           // 3) SUBIDA de req_id → congelar receta. NO publicar id_ok todavía.
           IF (#SupervisorCmdReqId AND NOT #L_IdEvalDone) THEN
               #Cfg_Pns := #SupervisorCmdPns;
               #Cfg_ReferencePart := #SupervisorCmdReferencePart;
               #Cfg_EndEffector := #SupervisorCmdEndEffector;
               #Cfg_UtTeach := #SupervisorCmdUtTech;
               #Cfg_TeachReq := #SupervisorCmdTeachReq;
               #Cfg_PaCheckReq := #SupervisorCmdPaCheckReq;
               #Cfg_TcgReq := #SupervisorCmdTcgReq;

               //4) Resuelve índices de programa por pieza (tu mapeo PIEZA1/2/3)
               IF #Cfg_ReferencePart = 'RefA400M' AND #Cfg_Pns ='M551B2810006-A01' THEN
                   //PART NUMBER QUE ME ENVIARÁ DE LA PIEZA SERÁ M551B2810006-A01 
                   //  REVESTIMIENTO INF IZQ - A400M
                   #PartProgIdx := 1;
                   #RefProgIdx := 1;
               ELSIF #Cfg_ReferencePart = 'RefF10X' AND #Cfg_Pns ='F46C551713119B01'   THEN
                   //PART NUMBER QUE ME ENVIARÁ SERÁ F46C551713110B01
                   //CARENA INF. IZQ HTP/VTP - Sandwich - FALCON
                   #PartProgIdx := 2;
                   #RefProgIdx := 2;
               ELSIF #Cfg_ReferencePart = 'RefEFA' AND #Cfg_Pns ='J57462100-406' THEN
                   #PartProgIdx := 3;
                   #RefProgIdx := 3;
               ELSE
                   #PartProgIdx := 100;
                   #RefProgIdx := 100;
               END_IF;

               #L_IdEvalDone := TRUE;
           END_IF;

           // 5) BAJADA de req_id → PUBLICAR id_ok y decidir salto.
           IF ((NOT #SupervisorCmdReqId) AND #L_IdEvalDone) THEN

               //5.1) Calcula PclstatusIdOk
               #PlcStatusIdOk :=
               ("PlcStatus".plcOk AND "SupervisorCmd".supervisorOk AND "PlcStatus".robotOk AND "PlcStatus".safetyOk
               AND "PlcStatus".airOk AND "PlcStatus".inspWaterOk AND "PlcStatus".tankWaterOk)
               AND (#Cfg_EndEffector >= 1) AND (#Cfg_EndEffector <= 5);

               #PlcStatusIdRunning := FALSE;

               //5.2)Decide siguiente STEP
               IF NOT #PlcStatusIdOk THEN
                   #PlcStatusStepPlc := #cSTEP_ID;
               ELSE
                   IF #Cfg_TeachReq THEN
                       #PlcStatusStepPlc := #cSTEP_TEACH;
                   ELSE
                       #PlcStatusStepPlc := #cSTEP_STARTUS;
                   END_IF;
               END_IF;

               #L_IdEvalDone := FALSE;
           END_IF;


           // ===============================================================
           // 2) TEACHING (pág. 4) — multi-PN: rearmar teach_ready por PN
           // FÍSICO: si la herramienta necesaria para teaching no está montada,
           // el KUKA cambia en Staübli al stand indicado (usa Supervisor.end-effector).
           // Luego, el KUKA se mueve al INICIO del PN siguiente y pone un bit de “en posición”.
           // Ese bit alimenta TeachAtStart=TRUE. Entonces EL PLC arma teach_ready (p. 4).
           // Repetir por cada PN mientras teach_app_running=TRUE.
           // ===============================================================
           (*  #cSTEP_TEACH:

             IF "SupervisorCmd".teachAppRunning THEN
                   IF (NOT "SupervisorCmd".teachRunning) AND TeachAtStart THEN
                       "PlcStatus".teachReady := TRUE;
                   END_IF;

                   IF "SupervisorCmd".teachRunning THEN
                       "PlcStatus".teachReady := FALSE;
                       teachWasRunning := TRUE;
                   END_IF;

                   // Fin de una trayectoria de teaching (sin abandonar la app)
                   IF (NOT "SupervisorCmd".teachRunning) AND teachWasRunning THEN
                       teachWasRunning := FALSE;
                   END_IF;

               ELSE
                   // Cierre de la app: salto según teach_state
                   IF "SupervisorCmd".teachState THEN
                       "PlcStatus".stepPlc := cSTEP_STARTUS;
                   ELSE
                       "PlcStatus".stepPlc := cSTEP_ID;
                   END_IF;
               END_IF;
           END_IF;*)




           // ===============================================================
           // 3) START US (pág. 5) — armar cuando “previous task done”
           // FÍSICO: KUKA AUT EXT cambia (si hace falta) al efector de INSPECCIÓN
           // requerido (Supervisor.end-effector, p. 1). Cuando:
           //   - Herramienta correcta acoplada (Staübli OK),
           //   - servicios/enclavamientos OK (safety/air/water/tank),
           //   - robot en posición segura para inicializar el UT,
           // el secuenciador pone StartUSReady=TRUE. El PLC arma start_us_ready.
           // Supervisor hace init UT (start_us_running/state_us). (p. 5)
           // ===============================================================
       #cSTEP_STARTUS:

           // Al entrar, ordena al robot cargar la herramienta decidida en ID
           IF #firstScan THEN
               #SupervisorCmdSeq := #SupervisorCmdSeq + 1;
               #WantCode_uint := #cKUKA_REQ_TOOL;
               #WantToolRequestId := (#Cfg_EndEffector);       // 1..5
           END_IF;

           // El PLC arma startUsReady SI el entorno/robot están listos y todavía no corre
           IF #StartUSReady AND (#WantCode_uint = 0) AND ("ToolInRobot_DB".toolInRobot_Num = #Cfg_EndEffector) AND NOT #SupervisorCmdStartUsRunning THEN
               #PlcStatusStartUsReady := TRUE;
           END_IF;

           // Cuando arranca, baja el "ready" y registra que realmente empezó
           IF #SupervisorCmdStartUsRunning THEN
               #PlcStatusStartUsReady := FALSE;
               #startUSWasRunning := TRUE;
           END_IF;

           // Al terminar: salto a PA o a Gain según lo congelado en ID
           IF (NOT #SupervisorCmdStartUsRunning)  AND #startUSWasRunning THEN
               #startUSWasRunning := FALSE;
               IF NOT #SupervisorCmdStateUs THEN
                   #PlcStatusStepPlc := #cSTEP_ID;
               ELSE
                   IF #Cfg_PaCheckReq THEN
                       #PlcStatusStepPlc := #cSTEP_PA_BAL;
                   ELSE
                       #PlcStatusStepPlc := #cSTEP_GAIN;
                   END_IF;
               END_IF;
           END_IF;


           // ===============================================================
           // 4) DEAD ELEMENT CHECK & BALANCING (pág. 6)
           //FÍSICO: KUKA va a la pieza Perspex de calibración y, cuando está en
           // [CORREGIDO] Lógica secuencial robusta, GOTO determinista y Retracción.
           // ===============================================================
       #cSTEP_PA_BAL:
           CASE #paBalSubStep OF
               0: // Inicialización y GOTO_PERSPEX
                   // [MEJORA] Siempre enviar comando GOTO en firstScan.
                   IF #firstScan THEN
                       #SupervisorCmdSeq := #SupervisorCmdSeq + 1;
                       #WantCode_uint := #cKUKA_GOTO_PERSPEX;
                   END_IF;
                   #paBalSubStep := 10;
               10: // Esperar Posición en Perspex     
                   // [MEJORA] Esperar posición Y canal libre (Race condition fix)
                   IF #kukaAtPerspexPos AND (#WantCode_uint = 0) THEN
                       #paBalSubStep := 20;
                   END_IF;
               20: // Ready for Dead Element Check     
                   IF NOT "SupervisorCmd".elemRunning THEN
                       "PlcStatus".paCheckReady := TRUE;
                   END_IF;
                   IF "SupervisorCmd".elemRunning THEN
                       "PlcStatus".paCheckReady := FALSE;
                       #paBalSubStep := 30;
                   END_IF;
               30: // Dead Element Check Running       
                   IF NOT "SupervisorCmd".elemRunning THEN
                       IF "SupervisorCmd".elemState THEN
                           #paBalSubStep := 40; // OK -> Balancing
                       ELSE
                           // KO -> Almacenar resultado y retraer
                           #tempNextStep := #cSTEP_ID;
                           #paBalSubStep := 60; // Ir a retracción
                       END_IF;
                   END_IF;
               40: // Ready for Balancing (Supervisor inicia automáticamente)        
                   IF "SupervisorCmd".balRunning THEN
                       #paBalSubStep := 50;
                   END_IF;
               50: // Balancing Running        
                   IF NOT "SupervisorCmd".balRunning THEN
                       // Determinar el siguiente paso
                       IF "SupervisorCmd".balState THEN
                           #tempNextStep := #cSTEP_GAIN; // OK
                       ELSE
                           #tempNextStep := #cSTEP_ID; // KO
                       END_IF;
                       #paBalSubStep := 60; // Proceder a retracción
                   END_IF;

                   // --- [MEJORA] LÓGICA DE RETRACCIÓN ESPECÍFICA ---
               60: // Ordenar RETRACT_PERSPEX
                   // [MEJORA] Esperar disponibilidad del despachador (Race condition fix)
                   IF (#WantCode_uint = 0) THEN
                       #SupervisorCmdSeq := #SupervisorCmdSeq + 1;
                       #WantCode_uint := #cKUKA_RETRACT_PERSPEX; // 101
                       #paBalSubStep := 70;
                   END_IF;

               70: // Esperar Fin de Retracción
                   // Robot terminó (WantCode_uint reseteado por el despachador)
                   IF (#WantCode_uint = 0) THEN
                       // Transición al paso almacenado
                       "PlcStatus".stepPlc := #tempNextStep;
                   END_IF;
           END_CASE;

           // ===============================================================
           // 5) GAIN ADJUSTMENT (pág. 7)
           // FÍSICO: KUKA se posiciona en la referencia para ganancia estática;
           // [CORREGIDO] Lógica secuencial robusta, GOTO determinista y Retracción.
           // ===============================================================
       #cSTEP_GAIN:

           CASE #gainSubStep OF
               0: // Inicialización y GOTO_GAIN
                   // [MEJORA] Siempre enviar comando GOTO en firstScan.
                   IF #firstScan THEN
                       #SupervisorCmdSeq := #SupervisorCmdSeq + 1;
                       #WantCode_uint := #cKUKA_GOTO_GAIN;
                   END_IF;
                   #gainSubStep := 10;

               10: // Esperar Posición en Gain    
                   // [MEJORA] Esperar posición Y canal libre (Race condition fix)
                   IF #kukaAtGainPos AND (#WantCode_uint = 0) THEN
                       #gainSubStep := 20;
                   END_IF;

               20: // Ready for Gain (Supervisor)    
                   IF NOT "SupervisorCmd".gainRunning THEN
                       "PlcStatus".gainReady := TRUE;
                   END_IF;

                   IF "SupervisorCmd".gainRunning THEN
                       "PlcStatus".gainReady := FALSE;
                       #gainSubStep := 30;
                   END_IF;

               30: // Gain Running
                   IF NOT "SupervisorCmd".gainRunning THEN
                       // Determinar siguiente paso
                       IF "SupervisorCmd".gainState THEN
                           IF #Cfg_TcgReq THEN
                               #tempNextStep := #cSTEP_TCG;
                           ELSE
                               #tempNextStep := #cSTEP_SCAN_REF;
                           END_IF;
                       ELSE
                           #tempNextStep := #cSTEP_ID; // KO        
                       END_IF;
                       #gainSubStep := 40; // Proceder a retracción
                   END_IF;

                   // --- [MEJORA] LÓGICA DE RETRACCIÓN ESPECÍFICA ---
               40: // Ordenar RETRACT_GAIN
                   // [MEJORA] Esperar disponibilidad del despachador (Race condition fix) 
                   IF (#WantCode_uint = 0) THEN
                       #SupervisorCmdSeq := #SupervisorCmdSeq + 1;
                       #WantCode_uint := #cKUKA_RETRACT_GAIN; // 102
                       #gainSubStep := 50;
                   END_IF;
               50: // Esperar Fin de Retracción         
                   IF (#WantCode_uint = 0) THEN
                       "PlcStatus".stepPlc := #tempNextStep;
                   END_IF;

           END_CASE;




           // ===============================================================
           // (6) TCG CHECK / ADJUSTMENT — pág. 8 (multiposición)
           // FÍSICO: KUKA recorre varias posiciones TCG. Para cada posición:
           // [CORREGIDO] Handshake Manager, GOTO determinista, Race Condition Fix y Retracción.
           // ===============================================================
       #cSTEP_TCG:

           // [MEJORA] Siempre ordenar el primer movimiento al entrar.    
           IF #firstScan THEN
               #SupervisorCmdSeq := #SupervisorCmdSeq + 1;
               #WantCode_uint := #cKUKA_GOTO_TCG;
               #WantIndex := (#tcgIndex); // Debería ser 1
               #waitingNextTCGPos := TRUE;
           END_IF;

           // Rearme de espera.
           // [MEJORA] Esperar a KUKA en posición Y que el canal esté libre (Race condition fix).
           IF #waitingNextTCGPos AND #kukaAtTCGPos AND (#WantCode_uint = 0) THEN
               #waitingNextTCGPos := FALSE;
           END_IF;

           // tcg_ready sólo si no mide, no esperamos pos, y el Handshake Manager está libre.
           IF (NOT "SupervisorCmd".tcgInProgress) AND (NOT #waitingNextTCGPos) AND (#handshakeStep = 0) THEN
               "PlcStatus".tcgReady := TRUE;
           ELSE
               // Asegurar que tcgReady baja si alguna condición falla (ej. Supervisor inicia medición)     
               "PlcStatus".tcgReady := FALSE;
           END_IF;

           // --- [MEJORA] Handshake Manager (4-way Acknowledge) - PDF Pág. 8 ---
           CASE #handshakeStep OF
               0: // IDLE: Esperar solicitud (Priorizadas)
                   // Solo aceptar si no estamos esperando movimiento ni midiendo
                   IF (NOT #waitingNextTCGPos) AND (NOT "SupervisorCmd".tcgInProgress) THEN
                       IF "SupervisorCmd".tcgNextStep THEN
                           #handshakeStep := 1; // NEXT
                       ELSIF "SupervisorCmd".reqRefPart THEN
                           #handshakeStep := 2; // ReqRefPart (Salida)
                       ELSIF "SupervisorCmd".reqStopCycle THEN
                           #handshakeStep := 3; // StopCycle (Salida)
                       ELSIF "SupervisorCmd".reqTcgAdj THEN
                           #handshakeStep := 4; // TcgAdj (Permanece en TCG) 
                       END_IF;
                   END_IF;

                   //1, 2, 3, 4: // SOLICITUD RECIBIDA: Enviar Acknowledge     
                   "PlcStatus".acknowledge := TRUE;
                   #handshakeStep := #handshakeStep + 10; // Pasar a esperar bajada
                   // --- Esperar Bajada de Solicitud ---    
               11: // NEXT    
                   IF NOT "SupervisorCmd".tcgNextStep THEN
                       "PlcStatus".acknowledge := FALSE;
                       // Acción NEXT: Pasar a esperar disponibilidad del canal antes de enviar.
                       #handshakeStep := 21;
                   END_IF;
               12: // ReqRefPart (Salida)
                   IF NOT "SupervisorCmd".reqRefPart THEN
                       "PlcStatus".acknowledge := FALSE;
                       // Acción: Preparar retracción antes de saltar.
                       #tempNextStep := #cSTEP_SCAN_REF;
                       #handshakeStep := 50; // Ir a retracción
                   END_IF;

               13: // StopCycle (Salida)     
                   IF NOT "SupervisorCmd".reqStopCycle THEN
                       "PlcStatus".acknowledge := FALSE;
                       // Acción: Preparar retracción antes de saltar. 
                       #tempNextStep := #cSTEP_ID;
                       #handshakeStep := 50; // Ir a retracción
                   END_IF;

               14: // TcgAdj (Permanece)     
                   IF NOT "SupervisorCmd".reqTcgAdj THEN
                       "PlcStatus".acknowledge := FALSE;
                       // Acción: Permanecer en TCG (Modo Ajuste).   
                       #handshakeStep := 0;
                   END_IF;

                   // --- Ejecución de NEXT (Sincronización con Despachador) ---
               21: // EJECUTAR NEXT (Wait for Dispatcher)
                   // [MEJORA] Evitar condición de carrera del despachador.
                   IF (#WantCode_uint = 0) THEN
                       // Canal libre -> Enviar comando GOTO_TCG
                       #tcgIndex := #tcgIndex + 1;
                       #SupervisorCmdSeq := #SupervisorCmdSeq + 1;
                       #WantCode_uint := #cKUKA_GOTO_TCG;
                       #WantIndex := (#tcgIndex);
                       #waitingNextTCGPos := TRUE;
                       #handshakeStep := 0;
                   END_IF;

                   // --- LÓGICA DE RETRACCIÓN ESPECÍFICA (Para salidas del paso TCG) ---        
               50: // Ordenar RETRACT_TCG
                   IF (#WantCode_uint = 0) THEN
                       #SupervisorCmdSeq := #SupervisorCmdSeq + 1;
                       #WantCode_uint := #cKUKA_RETRACT_TCG; // 103
                       #handshakeStep := 60;
                   END_IF;

               60: // Esperar Fin de Retracción      
                   IF (#WantCode_uint = 0) THEN
                       "PlcStatus".stepPlc := #tempNextStep; // Ir al paso almacenado
                       #handshakeStep := 0;
                   END_IF;
           END_CASE;



           // ===============================================================
           // (7) SCAN REFERENCE ACQUISITION — pág. 10
           // FÍSICO: KUKA carga PN/frame y se coloca en el punto de INICIO de
           // la trayectoria de referencia. Tu lógica pone AtRefScanStart=TRUE cuando
           // está en posición. 
           // // [MEJORA] GOTO determinista y Sincronización robusta.
           // ===============================================================
       #cSTEP_SCAN_REF:

           // Validación mínima de parámetros de scan que el PLC publica al Supervisor
           #validScanParams := (LEN("PlcStatus".idScan) > 0) AND ("PlcStatus".xSize > 0.0) AND ("PlcStatus".ySize > 0.0);

           // [MEJORA] Siempre enviar comando GOTO en firstScan.
           IF #firstScan THEN
               #SupervisorCmdSeq := #SupervisorCmdSeq + 1;
               #WantCode_uint := #cKUKA_GOTO_REF_START; // CASE 420
               #WantProgRequestId := (#RefProgIdx); // índice de programa REF por pieza
           END_IF;

           // Permiso de arranque
           // [MEJORA] Esperar posición Y canal libre antes de dar Ready.
           IF #kukaAtRefScanStartPos AND (#WantCode_uint = 0) AND #validScanParams AND NOT "SupervisorCmd".scanRefRunning THEN
               "PlcStatus".scanRefStart := TRUE;
           END_IF;

           // Cuando el Supervisor arranca → ejecutar trayectoria (CASE 432)
           IF (NOT #scanRefWasRunning) AND "SupervisorCmd".scanRefRunning THEN
               // [MEJORA] Esperar a que el despachador esté libre antes de enviar RUN.
               IF (#WantCode_uint = 0) THEN
                   #SupervisorCmdSeq := #SupervisorCmdSeq + 1;
                   #WantCode_uint := #cKUKA_RUN_REF_PATH;
                   #WantProgRequestId := (#RefProgIdx);
                   #scanRefWasRunning := TRUE; // Marcar como iniciado solo tras enviar comando
               END_IF;
           END_IF;

           IF "SupervisorCmd".scanRefRunning THEN
               // Bajar Ready cuando el robot termina físicamente  
               IF #kukaRefScanFinished THEN
                   "PlcStatus".scanRefStart := FALSE;
               END_IF;
           END_IF;

           // Fin del escaneo    
           IF (NOT "SupervisorCmd".scanRefRunning) AND #scanRefWasRunning THEN
               #scanRefWasRunning := FALSE;
               "PlcStatus".scanRefStart := FALSE;
               IF NOT "SupervisorCmd".scanRefState THEN
                   "PlcStatus".stepPlc := #cSTEP_ID;
               ELSE
                   "PlcStatus".stepPlc := #cSTEP_SCAN_INSP;
               END_IF;
           END_IF;


           // ===============================================================
           // (8) SCAN INSPECTION — pág. 11
           // FÍSICO: KUKA se coloca en INICIO de la(s) trayectoria(s) de inspección
           // [CORREGIDO] Handshake Manager, GOTO determinista y Sincronización robusta.
           // ===============================================================
       #cSTEP_SCAN_INSP:

           #validScanParams := (LEN("PlcStatus".idScan) > 0) AND ("PlcStatus".xSize > 0.0) AND ("PlcStatus".ySize > 0.0);

           // [MEJORA] Siempre enviar comando GOTO en firstScan.
           IF #firstScan THEN
               #SupervisorCmdSeq := #SupervisorCmdSeq + 1;
               #WantCode_uint := #cKUKA_GOTO_INSP_START;
               #WantProgRequestId := (#PartProgIdx);
           END_IF;

           // Permiso de arranque
           // [MEJORA] Esperar posición, canal libre y handshake libre antes de dar Ready.
           IF #kukaAtInspScanStartPos AND (#WantCode_uint = 0) AND #validScanParams AND NOT "SupervisorCmd".scanInsprunning AND (#handshakeStep = 0) THEN
               "PlcStatus".scanInspStart := TRUE;
           END_IF;

           // Al arrancar → ejecutar trayectoria (CASE 433)
           IF (NOT #scanInspWasRunning) AND "SupervisorCmd".scanInsprunning THEN
               // [MEJORA] Esperar a que el despachador esté libre antes de enviar RUN.
               IF (#WantCode_uint = 0) THEN
                   #SupervisorCmdSeq := #SupervisorCmdSeq + 1;
                   #WantCode_uint := #cKUKA_RUN_INSP_PATH;
                   #WantProgRequestId := (#PartProgIdx);
                   #scanInspWasRunning := TRUE; // Marcar como iniciado solo tras enviar comando
               END_IF;
           END_IF;


           IF "SupervisorCmd".scanInsprunning THEN
               // Bajar Ready cuando el robot termina físicamente
               IF #kukaInspScanFinished THEN
                   "PlcStatus".scanInspStart := FALSE;
               END_IF;
           END_IF;

           // Fin del escaneo 
           IF (NOT "SupervisorCmd".scanInsprunning) AND #scanInspWasRunning THEN
               #scanInspWasRunning := FALSE;
               "PlcStatus".scanInspStart := FALSE;

               IF NOT "SupervisorCmd".scanInspState THEN
                   "PlcStatus".stepPlc := #cSTEP_ID;
               ELSE
                   // Escaneo OK -> Activar Handshake Manager para esperar req_verif
                   #handshakeStep := 1;
               END_IF;
           END_IF;
           // [MEJORA] Handshake Manager (4-way) para req_verif (PDF Pág. 11)     
               CASE #handshakeStep OF
                   1: // Esperando req_verif
                       IF "SupervisorCmd".reqVerif THEN
                           #handshakeStep := 2;
                       END_IF;

                   2: // Enviar Acknowledge       
                       "PlcStatus".acknowledge := TRUE;
                       #handshakeStep := 3;

                   3: // Esperar bajada de req_verif    
                       IF NOT "SupervisorCmd".reqVerif THEN
                           "PlcStatus".acknowledge := FALSE;
                           // Acción: Saltar a Verificación 
                           "PlcStatus".stepPlc := #cSTEP_SCAN_REF_VERIF;
                           #handshakeStep := 0;
                       END_IF;
               END_CASE;





           // ===============================================================
           // (9) SCAN REFERENCE VERIFICATION — pág. 12
           // FÍSICO: KUKA vuelve al INICIO de la trayectoria de verificación de ref.
           // [CORREGIDO] Handshake Manager, Orden Faltante, GOTO y Sincronización.
           // ===============================================================
       #cSTEP_SCAN_REF_VERIF:

           #validScanParams := (LEN("PlcStatus".idScan) > 0) AND ("PlcStatus".xSize > 0.0) AND ("PlcStatus".ySize > 0.0);

           // [MEJORA] Siempre enviar comando GOTO en firstScan.
           IF #firstScan THEN
               #SupervisorCmdSeq := #SupervisorCmdSeq + 1;
               #WantCode_uint := #cKUKA_GOTO_REF_START;
               #WantProgRequestId := (#RefProgIdx);
           END_IF;
           // Permiso de arranque    
           // [MEJORA] Esperar posición, canal libre y handshake libre antes de dar Ready.
           IF #kukaAtRefScanStartPos AND (#WantCode_uint = 0) AND #validScanParams AND NOT "SupervisorCmd".scanRefRunning AND (#handshakeStep = 0) THEN
               "PlcStatus".scanRefStart := TRUE;
           END_IF;

           // [CORRECCIÓN] Al arrancar -> ejecutar trayectoria (Faltaba esta orden)
           IF (NOT #scanRefWasRunning) AND "SupervisorCmd".scanRefRunning THEN
               // [MEJORA] Esperar a que el despachador esté libre antes de enviar RUN.
               IF (#WantCode_uint = 0) THEN
                   #SupervisorCmdSeq := #SupervisorCmdSeq + 1;
                   #WantCode_uint := #cKUKA_RUN_REF_PATH; // 432
                   #WantProgRequestId := (#RefProgIdx);
                   #scanRefWasRunning := TRUE; // Marcar como iniciado solo tras enviar comando
               END_IF;
           END_IF;

           IF "SupervisorCmd".scanRefRunning THEN
               // [CORRECCIÓN] Bajar scanRefStart cuando el robot termina (PDF p.12).
               IF #kukaRefScanFinished THEN
                   "PlcStatus".scanRefStart := FALSE;
               END_IF;
           END_IF;

           // Fin del escaneo de verificación
           IF (NOT "SupervisorCmd".scanRefRunning) AND #scanRefWasRunning THEN
               #scanRefWasRunning := FALSE;
               "PlcStatus".scanRefStart := FALSE;
               IF NOT "SupervisorCmd".scanRefState THEN
                   "PlcStatus".stepPlc := #cSTEP_ID;
               ELSE
                   // OK -> Activar Handshake Manager para esperar decisiones    
                   #handshakeStep := 1;
               END_IF;
           END_IF;

           // [MEJORA] Handshake Manager (4-way) (PDF Pág. 12)
           CASE #handshakeStep OF
               1: // Esperando decisiones (Priorizadas)
                   IF "SupervisorCmd".reqPreEval THEN
                       #handshakeStep := 2; // Pre-eval
                   ELSIF "SupervisorCmd".reqIdentificationState THEN
                       #handshakeStep := 3; // Nuevo ciclo
                   END_IF;
                   // 2, 3: // Enviar Acknowledge
                   "PlcStatus".acknowledge := TRUE;
                   #handshakeStep := #handshakeStep + 10;
               12: // Esperar bajada (Pre-eval)     
                   IF NOT "SupervisorCmd".reqPreEval THEN
                       "PlcStatus".acknowledge := FALSE;
                       "PlcStatus".stepPlc := #cSTEP_PRE_EVAL;
                       #handshakeStep := 0;
                   END_IF;

               13: // Esperar bajada (Nuevo Ciclo)      
                   IF NOT "SupervisorCmd".reqIdentificationState THEN
                       "PlcStatus".acknowledge := FALSE;
                       // Nota: No se requiere GOTO_SAFE aquí, ya que el escaneo no es peligroso.
                       "PlcStatus".stepPlc := #cSTEP_ID;
                       #handshakeStep := 0;
                   END_IF;
           END_CASE;

           // ===============================================================
           // (10) PRE‑EVALUATION / MARKING — pág. 13
           // FÍSICO: si la herramienta de marcado no está montada, el KUKA cambia
           // en Staübli al stand de “marking” según requiera el proceso; tras estar
           // [CORREGIDO] Gestión de herramienta, ejecución física, Handshake y movimiento seguro.
           // ===============================================================
       #cSTEP_PRE_EVAL:

           // --- [MEJORA] Handshake Manager (4-way) para Nuevo ciclo + GOTO_SAFE ---  
           CASE #handshakeStep OF
               0: // Idle: Esperar solicitud de nuevo ciclo       
                   // Solo permitir si el marcado no está en curso   
                   IF "SupervisorCmd".reqIdentificationState AND (NOT "PlcStatus".markRunning) THEN
                       #handshakeStep := 1;
                   END_IF;
               1: // Enviar Ack    
                   "PlcStatus".acknowledge := TRUE;
                   #handshakeStep := 2;
               2: // Esperar bajada de la solicitud
                   IF NOT "SupervisorCmd".reqIdentificationState THEN
                       "PlcStatus".acknowledge := FALSE;
                       // Acción: Preparar para ir a Safe antes de ID    
                       #handshakeStep := 3;
                   END_IF;

                   // [MEJORA] Mover a Safe antes de saltar a ID      
               3: // Enviar GOTO_SAFE (Esperar disponibilidad del despachador)   
                   IF (#WantCode_uint = 0) THEN
                       #SupervisorCmdSeq := #SupervisorCmdSeq + 1;
                       //#WantCode_uint := #cKUKA_GOTO_SAFE; // 100
                       #handshakeStep := 4;
                   END_IF;

               4: // Esperar fin de GOTO_SAFE
                   IF (#WantCode_uint = 0) THEN
                       // Llegó a Safe -> Saltar a ID
                       "PlcStatus".stepPlc := #cSTEP_ID;
                       #handshakeStep := 0;
                   END_IF;
           END_CASE;

           // --- [MEJORA] Máquina de estados de Marcado ---
           CASE #markingSubStep OF
               0: // Inicialización (Al entrar al paso)
                   #markingSubStep := 10;
               10: // Cambio de Herramienta (a Marcador)     
                   // Solo si no la tiene ya y los canales están libres
                   IF ("ToolInRobot_DB".toolInRobot_Num <> 3) AND (#WantCode_uint = 0) AND (#handshakeStep = 0) THEN
                       #SupervisorCmdSeq := #SupervisorCmdSeq + 1;
                       #WantCode_uint := #cKUKA_REQ_TOOL;
                       #WantToolRequestId := #cTOOL_MARKER;
                   END_IF;

                   // Transición cuando tenga la herramienta y el canal esté libre    
                   IF ("ToolInRobot_DB".toolInRobot_Num = #cTOOL_MARKER) AND (#WantCode_uint = 0) THEN
                       #markingSubStep := 20;
                   END_IF;

               20: // Esperar Petición de Marcado (reqMark)
                   // Solo si el handshake general está libre
                   IF "SupervisorCmd".reqMark AND (#handshakeStep = 0) THEN
                       // 1. Transferir coordenadas al buffer (Asume Supervisor.pointCoordinates es ARRAY[0..5] OF REAL)
                       // #WantMarkCoords[0] := "SupervisorCmd".pointCoordinates[0]; // X
                       // ... (Copiar Y, Z, A, B, C) ...
                       // 2. Preparar estado y pasar a envío de comando
                       "PlcStatus".markState := FALSE;
                       "PlcStatus".markRunning := TRUE;
                       #markingSubStep := 30;
                   END_IF;

               30: // Enviar Comando al Robot (Esperar disponibilidad)    
                   // [MEJORA] Esperar a que el despachador esté libre.
                   IF (#WantCode_uint = 0) THEN
                       #SupervisorCmdSeq := #SupervisorCmdSeq + 1;
                       #WantCode_uint := #cKUKA_MARK_POINT; // Código 501
                       #markingSubStep := 40;
                   END_IF;

               40: // Ejecución en Progreso (Esperar fin en KUKA)  
                   // Esperar a que el robot termine el comando (WantCode_uint vuelve a 0)
                   IF (#WantCode_uint = 0) THEN
                       // El marcado ha terminado físicamente.
                       "PlcStatus".markState := #MarkingDone; // Leer resultado físico
                       #markingSubStep := 50;
                   END_IF;

               50: // Finalizado (Esperar que Supervisor baje reqMark - PDF p.13)
                   IF NOT "SupervisorCmd".reqMark THEN
                       "PlcStatus".markRunning := FALSE;
                       "PlcStatus".markRunning := FALSE;
                   END_IF;

           END_CASE;
       ELSE
           "PlcStatus".stepPlc := #cSTEP_ID;

   END_CASE;


   // ---------------------------------------------------------------
   // [2] DESPACHO AL KUKA (toggle goTrigger cuando el canal esté libre)
   //     • Este bloque “consume” el slot WantCmd → publica parámetros
   //       en los registros PNIO (con SWAP) → toggle de goTrigger.
   //     • El robot deberá igualar rbDone := goTrigger al terminar.
   // ---------------------------------------------------------------

   CASE #state OF
       0: // IDLE -> GO == ACK

           // "cancelGo" := FALSE;

           IF (#SupervisorCmdSeq <> #lastSeq) THEN

               IF  "goTrigger" = "rbDone" THEN

                   #code_int := #WantCode_uint;  // “code_int” que viajará al KRC

                   // (Códigos existentes 201, 414, 420, 432, 421, 433 se mantienen igual)

                   IF #code_int = 201 THEN
                       // id de herramienta → WORD+SWAP
                       // #Cfg_EndEffector
                       #toolReqId := SWAP(INT_TO_WORD(#WantToolRequestId));

                   END_IF;

                   IF #code_int = 414 THEN  //GOTO_TCG
                       // id de herramienta → WORD+SWAP
                       "requestIndexKuka" := SWAP(UINT_TO_WORD(#WantIndex));

                   END_IF;

                   IF #code_int = 420 THEN // GOTO_REF_START
                       // id de herramienta → WORD+SWAP
                       "programReqId" := SWAP(UINT_TO_WORD(#WantProgRequestId));

                   END_IF;

                   IF #code_int = 432 THEN // RUN_REF_PATH
                       // id de herramienta → WORD+SWAP
                       "programReqId" := SWAP(UINT_TO_WORD(#WantProgRequestId));

                   END_IF;

                   IF #code_int = 421 THEN // GOTO_REF_START
                       // id de herramienta → WORD+SWAP
                       "programReqId" := SWAP(UINT_TO_WORD(#WantProgRequestId));

                   END_IF;

                   IF #code_int = 433 THEN // RUN_INSP_PATH

                       "programReqId" := SWAP(UINT_TO_WORD(#WantProgRequestId));

                   END_IF;

                   // [MEJORA] Transferencia de Coordenadas para Marcado (501)
                  // IF #code_int = #cKUKA_MARK_POINT THEN
                        // Convertir REAL a DWORD/DINT y hacer SWAP para enviar por Profinet
                        //  // Ejemplo: "ProfinetOutputs".MarkX := SWAP(REAL_TO_DWORD(#WantMarkCoords[0]));
                   //END_IF;

                   // 2) Publicar código de movimiento
                   #moveCodeKuka := SWAP(UINT_TO_WORD(#code_int));   // KRC leerá "MoveCode" = INT

                   // 3) Disparo del GO: toggle de goTrigger (rbDone ≠ goTrigger → pedido activo)
                   "goTrigger" := NOT "goTrigger";

                   #lastSeq := #SupervisorCmdSeq;          // <-- memoriza!
                   #state := 20;

               END_IF;
           END_IF;

       20: // BUSY

           //#code_int := #KukaControlCmdCode;

           // CANCEL pedido en BUSY → avisar al KRC y ACK de la ORDEN ACTIVA
           IF #code_int = 903 THEN
               "cancelGo" := TRUE;
           END_IF;

           // Fin normal (o tras el cancel, cuando KRC cierra el canal por nivel)

           IF ("rbDone" = "goTrigger") THEN
               // 4) Vaciar slot de pendiente
               #WantCode_uint := 0;
               #WantProgRequestId := 0;
               #WantToolRequestId := 0;
               #WantIndex := 0;
               #state := 0;                            // vuelve a IDLE
           END_IF;

   END_CASE;
END_REGION
END_FUNCTION_BLOCK

ORGANIZATION_BLOCK "Main"   // OB1, LAD, ProgramCycle
TITLE = "Main Program Sweep (Cycle)"
{ S7_Optimized_Access := 'TRUE' }
VERSION : 0.1
   VAR_INPUT
      Initial_Call : Bool;   // Initial call of this OB
      Remanence : Bool;   // =True, if remanent data are available
   END_VAR
   VAR_TEMP
      evtEnterSrv : Bool;   // // Eventos de modo service jog
      evtEnterAuto : Bool;   // // Eventos de modo auto
      muxSelStb : Bool;
      muxStartStb : Bool;
      muxPgno : Byte;
      u : UDInt;
   END_VAR
BEGIN

REGION Network 1 (SCL): // ====================== REANUDAR MOVIMIENTO AUTOMATICO EXTERNO ======================
   // // —— Enlaza estos símbolos a tus %I en el árbol de dispositivos ——
   //   // EStop_DI, SafeDoor_DI, AirPressure_DI, WaterInsp_DI, WaterTank_DI, RobotReady_DI, ...
   "$MOVE_ENABLE" := TRUE;
   "$I_O_ACT" := TRUE;
   //"$DRIVES_OFF" := FALSE;

   "PlcStatus".systemArmed := FALSE;
   "PlcStatus".robotInAutExt := "$EXT";
   "PlcStatus".robotInHome := "$IN_HOME";
END_REGION

REGION Network 2: REANUDAR MOVIMIENTO EN KUKA
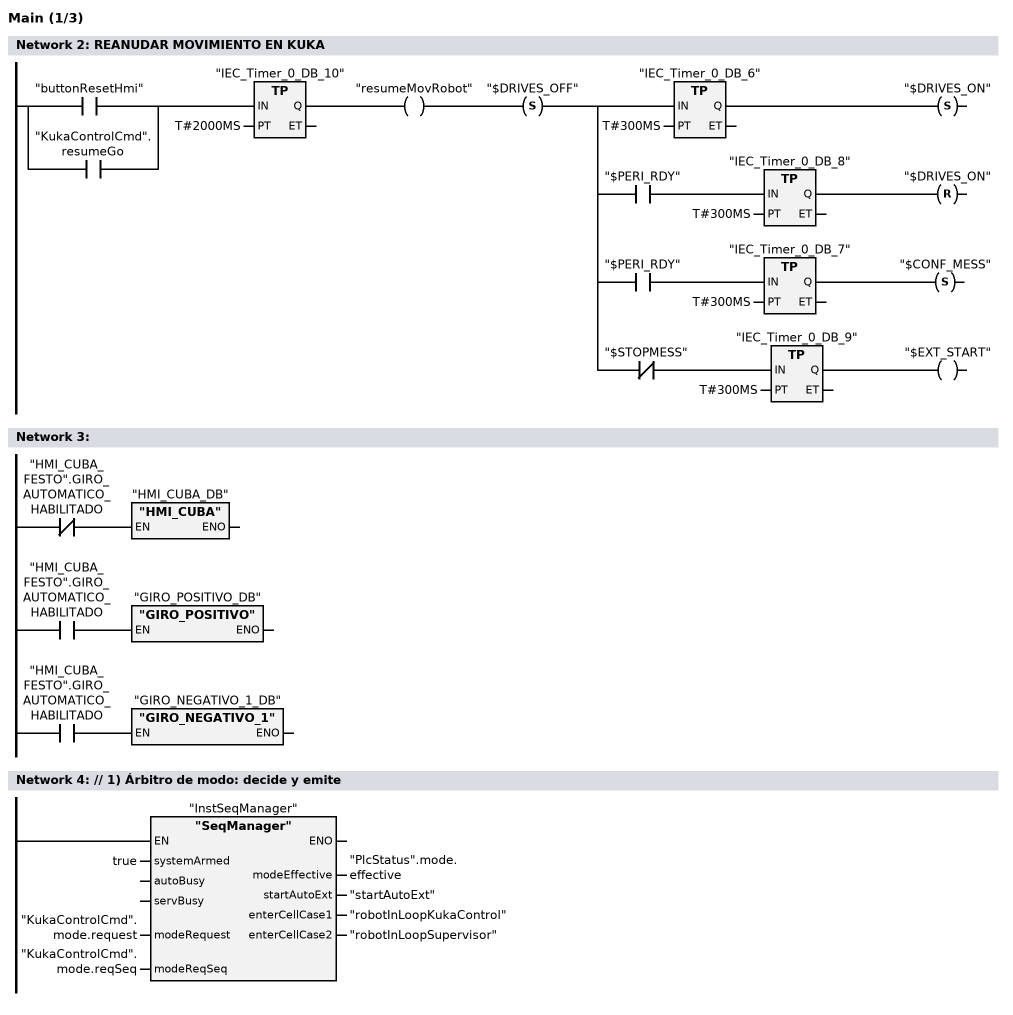
   "IEC_Timer_0_DB_10".TP(IN := "buttonResetHmi" OR "KukaControlCmd".resumeGo, PT := T#2000MS);
   "resumeMovRobot" := "IEC_Timer_0_DB_10".Q;
   IF "IEC_Timer_0_DB_10".Q THEN "$DRIVES_OFF" := TRUE; END_IF;
   "IEC_Timer_0_DB_6".TP(IN := "IEC_Timer_0_DB_10".Q, PT := T#300MS);
   IF "IEC_Timer_0_DB_6".Q THEN "$DRIVES_ON" := TRUE; END_IF;
   "IEC_Timer_0_DB_8".TP(IN := "IEC_Timer_0_DB_10".Q AND "$PERI_RDY", PT := T#300MS);
   IF "IEC_Timer_0_DB_8".Q THEN "$DRIVES_ON" := FALSE; END_IF;
   "IEC_Timer_0_DB_7".TP(IN := "IEC_Timer_0_DB_10".Q AND "$PERI_RDY", PT := T#300MS);
   IF "IEC_Timer_0_DB_7".Q THEN "$CONF_MESS" := TRUE; END_IF;
   "IEC_Timer_0_DB_9".TP(IN := "IEC_Timer_0_DB_10".Q AND NOT "$STOPMESS", PT := T#300MS);
   "$EXT_START" := "IEC_Timer_0_DB_9".Q;
END_REGION

REGION Network 3
   RUNG wire#powerrail
      I_Contact( "HMI_CUBA_FESTO".GIRO_AUTOMATICO_HABILITADO )
      "HMI_CUBA_DB"()
   END_RUNG
   RUNG wire#powerrail
      Contact( "HMI_CUBA_FESTO".GIRO_AUTOMATICO_HABILITADO )
      "GIRO_POSITIVO_DB"()
   END_RUNG
   RUNG wire#powerrail
      Contact( "HMI_CUBA_FESTO".GIRO_AUTOMATICO_HABILITADO )
      "GIRO_NEGATIVO_1_DB"()
   END_RUNG
   // the same network as SCL:
   IF NOT "HMI_CUBA_FESTO".GIRO_AUTOMATICO_HABILITADO THEN
       "HMI_CUBA_DB"();   // "HMI_CUBA"
   END_IF;
   IF "HMI_CUBA_FESTO".GIRO_AUTOMATICO_HABILITADO THEN
       "GIRO_POSITIVO_DB"();   // "GIRO_POSITIVO"
   END_IF;
   IF "HMI_CUBA_FESTO".GIRO_AUTOMATICO_HABILITADO THEN
       "GIRO_NEGATIVO_1_DB"();   // "GIRO_NEGATIVO_1"
   END_IF;
END_REGION

REGION Network 4: // 1) Árbitro de modo: decide y emite
   RUNG wire#powerrail
      "InstSeqManager"(systemArmed := true, autoBusy :=, servBusy :=, modeRequest := "KukaControlCmd".mode.request, modeReqSeq := "KukaControlCmd".mode.reqSeq, modeEffective => "PlcStatus".mode.effective, startAutoExt => "startAutoExt", enterCellCase1 => "robotInLoopKukaControl", enterCellCase2 => "robotInLoopSupervisor")
   END_RUNG
   // the same network as SCL:
   "InstSeqManager"(systemArmed := true,   // "SeqManager"
                    modeRequest := "KukaControlCmd".mode.request,
                    modeReqSeq := "KukaControlCmd".mode.reqSeq,
                    modeEffective => "PlcStatus".mode.effective,
                    startAutoExt => "startAutoExt",
                    enterCellCase1 => "robotInLoopKukaControl",
                    enterCellCase2 => "robotInLoopSupervisor");
END_REGION

REGION Network 5
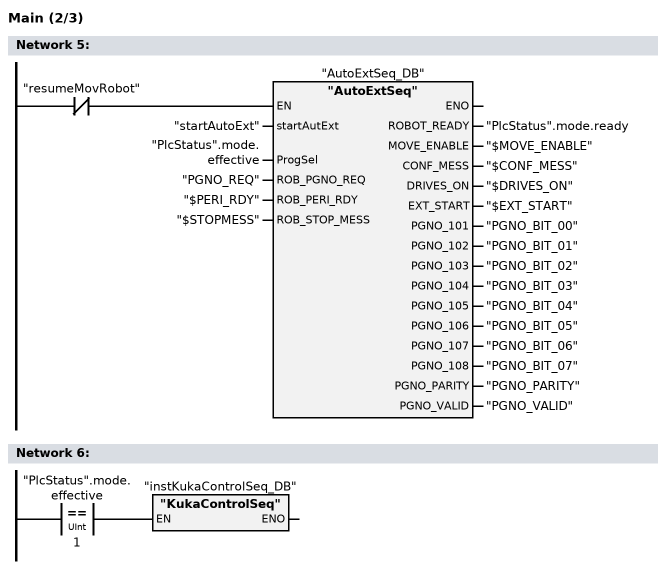
   RUNG wire#powerrail
      I_Contact( "resumeMovRobot" )
      "AutoExtSeq_DB"(startAutExt := "startAutoExt", ProgSel := "PlcStatus".mode.effective, ROB_PGNO_REQ := "PGNO_REQ", ROB_PERI_RDY := "$PERI_RDY", ROB_STOP_MESS := "$STOPMESS", ROBOT_READY => "PlcStatus".mode.ready, MOVE_ENABLE => "$MOVE_ENABLE", CONF_MESS => "$CONF_MESS", DRIVES_ON => "$DRIVES_ON", EXT_START => "$EXT_START", PGNO_101 => "PGNO_BIT_00", PGNO_102 => "PGNO_BIT_01", PGNO_103 => "PGNO_BIT_02", PGNO_104 => "PGNO_BIT_03", PGNO_105 => "PGNO_BIT_04", PGNO_106 => "PGNO_BIT_05", PGNO_107 => "PGNO_BIT_06", PGNO_108 => "PGNO_BIT_07", PGNO_PARITY => "PGNO_PARITY", PGNO_VALID => "PGNO_VALID")
   END_RUNG
   // the same network as SCL:
   IF NOT "resumeMovRobot" THEN
       "AutoExtSeq_DB"(startAutExt := "startAutoExt",   // "AutoExtSeq"
                       ProgSel := "PlcStatus".mode.effective,
                       ROB_PGNO_REQ := "PGNO_REQ",
                       ROB_PERI_RDY := "$PERI_RDY",
                       ROB_STOP_MESS := "$STOPMESS",
                       ROBOT_READY => "PlcStatus".mode.ready,
                       MOVE_ENABLE => "$MOVE_ENABLE",
                       CONF_MESS => "$CONF_MESS",
                       DRIVES_ON => "$DRIVES_ON",
                       EXT_START => "$EXT_START",
                       PGNO_101 => "PGNO_BIT_00",
                       PGNO_102 => "PGNO_BIT_01",
                       PGNO_103 => "PGNO_BIT_02",
                       PGNO_104 => "PGNO_BIT_03",
                       PGNO_105 => "PGNO_BIT_04",
                       PGNO_106 => "PGNO_BIT_05",
                       PGNO_107 => "PGNO_BIT_06",
                       PGNO_108 => "PGNO_BIT_07",
                       PGNO_PARITY => "PGNO_PARITY",
                       PGNO_VALID => "PGNO_VALID");
   END_IF;
END_REGION

REGION Network 6
   RUNG wire#powerrail
      { S7_Templates := "SrcType := UInt" } EQ_Contact(in1 := "PlcStatus".mode.effective, in2 := 1)
      "instKukaControlSeq_DB"()
   END_RUNG
   // the same network as SCL:
   IF "PlcStatus".mode.effective = 1 THEN
       "instKukaControlSeq_DB"();   // "KukaControlSeq"
   END_IF;
END_REGION

REGION Network 7
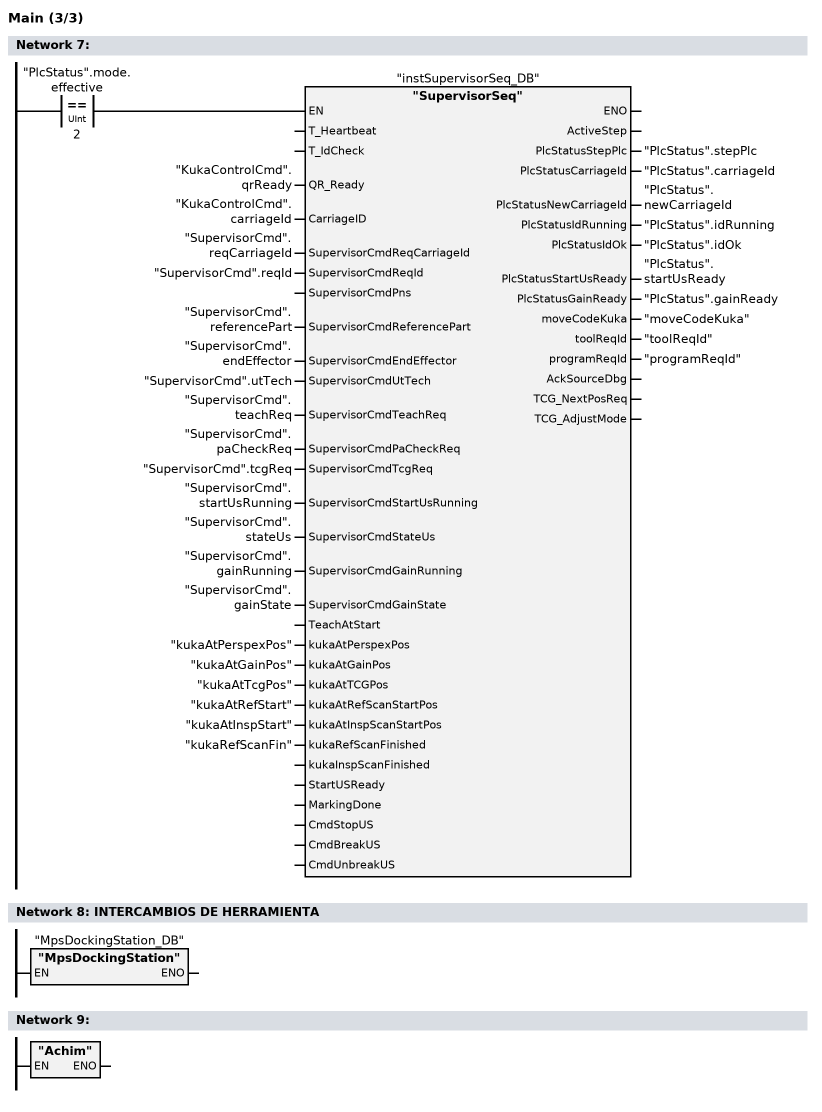
   RUNG wire#powerrail
      { S7_Templates := "SrcType := UInt" } EQ_Contact(in1 := "PlcStatus".mode.effective, in2 := 2)
      "instSupervisorSeq_DB"(T_Heartbeat :=, T_IdCheck :=, QR_Ready := "KukaControlCmd".qrReady, CarriageID := "KukaControlCmd".carriageId, SupervisorCmdReqCarriageId := "SupervisorCmd".reqCarriageId, SupervisorCmdReqId := "SupervisorCmd".reqId, SupervisorCmdPns :=, SupervisorCmdReferencePart := "SupervisorCmd".referencePart, SupervisorCmdEndEffector := "SupervisorCmd".endEffector, SupervisorCmdUtTech := "SupervisorCmd".utTech, SupervisorCmdTeachReq := "SupervisorCmd".teachReq, SupervisorCmdPaCheckReq := "SupervisorCmd".paCheckReq, SupervisorCmdTcgReq := "SupervisorCmd".tcgReq, SupervisorCmdStartUsRunning := "SupervisorCmd".startUsRunning, SupervisorCmdStateUs := "SupervisorCmd".stateUs, SupervisorCmdGainRunning := "SupervisorCmd".gainRunning, SupervisorCmdGainState := "SupervisorCmd".gainState, TeachAtStart :=, kukaAtPerspexPos := "kukaAtPerspexPos", kukaAtGainPos := "kukaAtGainPos", kukaAtTCGPos := "kukaAtTcgPos", kukaAtRefScanStartPos := "kukaAtRefStart", kukaAtInspScanStartPos := "kukaAtInspStart", kukaRefScanFinished := "kukaRefScanFin", kukaInspScanFinished :=, StartUSReady :=, MarkingDone :=, CmdStopUS :=, CmdBreakUS :=, CmdUnbreakUS :=, ActiveStep =>, PlcStatusStepPlc => "PlcStatus".stepPlc, PlcStatusCarriageId => "PlcStatus".carriageId, PlcStatusNewCarriageId => "PlcStatus".newCarriageId, PlcStatusIdRunning => "PlcStatus".idRunning, PlcStatusIdOk => "PlcStatus".idOk, PlcStatusStartUsReady => "PlcStatus".startUsReady, PlcStatusGainReady => "PlcStatus".gainReady, moveCodeKuka => "moveCodeKuka", toolReqId => "toolReqId", programReqId => "programReqId", AckSourceDbg =>, TCG_NextPosReq =>, TCG_AdjustMode =>)
   END_RUNG
   // the same network as SCL:
   IF "PlcStatus".mode.effective = 2 THEN
       "instSupervisorSeq_DB"(QR_Ready := "KukaControlCmd".qrReady,   // "SupervisorSeq"
                              CarriageID := "KukaControlCmd".carriageId,
                              SupervisorCmdReqCarriageId := "SupervisorCmd".reqCarriageId,
                              SupervisorCmdReqId := "SupervisorCmd".reqId,
                              SupervisorCmdReferencePart := "SupervisorCmd".referencePart,
                              SupervisorCmdEndEffector := "SupervisorCmd".endEffector,
                              SupervisorCmdUtTech := "SupervisorCmd".utTech,
                              SupervisorCmdTeachReq := "SupervisorCmd".teachReq,
                              SupervisorCmdPaCheckReq := "SupervisorCmd".paCheckReq,
                              SupervisorCmdTcgReq := "SupervisorCmd".tcgReq,
                              SupervisorCmdStartUsRunning := "SupervisorCmd".startUsRunning,
                              SupervisorCmdStateUs := "SupervisorCmd".stateUs,
                              SupervisorCmdGainRunning := "SupervisorCmd".gainRunning,
                              SupervisorCmdGainState := "SupervisorCmd".gainState,
                              kukaAtPerspexPos := "kukaAtPerspexPos",
                              kukaAtGainPos := "kukaAtGainPos",
                              kukaAtTCGPos := "kukaAtTcgPos",
                              kukaAtRefScanStartPos := "kukaAtRefStart",
                              kukaAtInspScanStartPos := "kukaAtInspStart",
                              kukaRefScanFinished := "kukaRefScanFin",
                              PlcStatusStepPlc => "PlcStatus".stepPlc,
                              PlcStatusCarriageId => "PlcStatus".carriageId,
                              PlcStatusNewCarriageId => "PlcStatus".newCarriageId,
                              PlcStatusIdRunning => "PlcStatus".idRunning,
                              PlcStatusIdOk => "PlcStatus".idOk,
                              PlcStatusStartUsReady => "PlcStatus".startUsReady,
                              PlcStatusGainReady => "PlcStatus".gainReady,
                              moveCodeKuka => "moveCodeKuka",
                              toolReqId => "toolReqId",
                              programReqId => "programReqId");
   END_IF;
END_REGION

REGION Network 8: INTERCAMBIOS DE HERRAMIENTA
   RUNG wire#powerrail
      "MpsDockingStation_DB"()
   END_RUNG
   // the same network as SCL:
   "MpsDockingStation_DB"();   // "MpsDockingStation"
END_REGION

REGION Network 9
   RUNG wire#powerrail
      "Achim"()
   END_RUNG
   // the same network as SCL:
   "Achim"();
END_REGION
END_ORGANIZATION_BLOCK

// folder: 20. Robot Services/AutoExt

FUNCTION_BLOCK "AutoExtSeq"   // FB31, LAD
{ S7_Optimized_Access := 'TRUE' }
VERSION : 0.1
   VAR_INPUT
      startAutExt : Bool;   // // Flanco para ejecutar CASE 1
      ProgSel : UInt;
      ROB_PGNO_REQ : Bool;
      ROB_PERI_RDY : Bool;
      ROB_STOP_MESS : Bool;
   END_VAR
   VAR_OUTPUT
      ROBOT_READY : Bool;
      MOVE_ENABLE : Bool := TRUE;
      CONF_MESS : Bool;
      DRIVES_ON : Bool;
      EXT_START : Bool;
      PGNO_101 : Bool;
      PGNO_102 : Bool;
      PGNO_103 : Bool;
      PGNO_104 : Bool;
      PGNO_105 : Bool;
      PGNO_106 : Bool;
      PGNO_107 : Bool;
      PGNO_108 : Bool;
      PGNO_PARITY : Bool;
      PGNO_VALID : Bool;
   END_VAR
   VAR
      "step" : Int;   // secuencia simple
      rStart : R_TRIG;
      rPgnoReq : R_TRIG;
      fPgnoReq : F_TRIG;
      tpConf : TP_TIME;
      tpDrives : TP_TIME;
      tpStart : TP_TIME;
      tpStartInit : TP_TIME;
      tStable : TON_TIME;
      pulseTime : Time := T#120ms;
      drivesPulse : Time := T#120ms;
      stableTime : Time := T#36ms;
      initStartPulse : Time := T#150ms;
      pgnoLatched : UInt;
      tPump : TP_TIME;
   END_VAR
BEGIN

REGION Network 1 (SCL): // === Secuencia Aut Ext ===
   /// 1) Detectores de flanco: se ejecutan SIEMPRE (cada ciclo de scan del plc)
   #rStart(CLK := #startAutExt);       // flanco de arranque de la secuencia
   #rPgnoReq(CLK := #ROB_PGNO_REQ);    // flanco de subida del PGNO_REQ
   #fPgnoReq(CLK := #ROB_PGNO_REQ);     // flanco de bajada del PGNO_REQ

   // ------------------------------ Máquina de estados ---------------------
   CASE #step OF

       0:   // IDLE: esperar flanco de arranque externo (#startAutExt 0→1)
           // No imprescindible, pero dejamos los temporizadores “quietos”
           #tpStartInit(IN := FALSE,
                        PT := #initStartPulse);
           #tpDrives(IN := FALSE,
                     PT := #initStartPulse);
           #tpStart(IN := FALSE,
                    PT := #initStartPulse);

           // Por defecto, PGNO inválido en reposo  para iniciar “limpio”
           #PGNO_VALID := FALSE;

           // Poner a '0' los bits PGNO mientras no haya petición del KRC
           #PGNO_101 := FALSE;
           #PGNO_102 := FALSE;
           #PGNO_103 := FALSE;
           #PGNO_104 := FALSE;
           #PGNO_105 := FALSE;
           #PGNO_106 := FALSE;
           #PGNO_107 := FALSE;
           #PGNO_108 := FALSE;
           #PGNO_PARITY := FALSE;


           // Arrancar SOLO en flanco de #startAutExt
           IF #rStart.Q THEN // SOLO en el flanco  (un ciclo)

               #ROBOT_READY := FALSE;   // el modo no está listo mientras arranca
               #step := 1;               // → primer pulso: DRIVES_ON
           END_IF;


       1:  // Pulso de DRIVES_ON (una sola vez por ciclo de autoext)
           // Llamamos al TP solo en este paso ⇒ genera un único pulso de ancho #drivesPulse
           #tpDrives(IN := TRUE,
                     PT := #drivesPulse);
           #DRIVES_ON := #tpDrives.Q;
           IF NOT #tpDrives.Q THEN
               #step := 2;          // cuando cae el pulso → segundo pulso
           END_IF;


       2:  // Pulso de CONF_MESS (también una sola vez)
           #tpConf(IN := TRUE,
                   PT := #drivesPulse);   // o #confPulse si quieres ancho distinto
           #CONF_MESS := #tpConf.Q;
           IF NOT #tpConf.Q THEN
               #step := 5;           // luego hacemos el pre‑start (salir de INIT)
           END_IF;


       5:  // PRE‑START: salir de AUTOEXT INIT con un start corto
           #tpStartInit(IN := TRUE,
                        PT := #initStartPulse);
           #EXT_START := #tpStartInit.Q;
           IF NOT #tpStartInit.Q THEN
               #step := 10; // → esperar petición de PGNO por parte del KRC
           END_IF;